			UConveyorIO.xExitBarCylinderRetract2:=0;
			iStep:=0;
		END_IF;
	END_CASE;
3:(*上料到出口*)
	CASE iStep OF
	0:(*各种初始化，能自动去3*)
		ConveyorIODown.xLoad:=0;
		ConveyorIOleft.xLoad:=0;
		ConveyorIORight.xLoad:=0;
		ConveyorIODown.xUnload:=0;
		ConveyorIOLeft.xUnload:=0;
		ConveyorIORight.xUnload:=0;
		UConveyorIO.xBatteryError:=0;
		UConveyorIO.xExitBarCylinderRetract1:=0;
		UConveyorIO.xExitBarCylinderRetract2:=0;
		ConveyorIODown.xPutInto:=0;
		ConveyorIOLeft.xPutInto:=0;
		ConveyorIORight.xPutInto:=0;
		IF m_xStep0 AND  ConveyorIODown.xEmpty THEN
			iStep:=1;
		ELSIF m_xStep0 AND NOT ConveyorIODown.xEmpty THEN
			iStep:=3;
		END_IF;	
	1:(*右顶升动作，等load*)
		IF UConveyorIO.xLiftCylinderExtendInit2 THEN
			UConveyorIO.xLiftCylinderExtend2:=0;
			UConveyorIO.xLiftCylinderRetract2:=1;
		ELSE
			UConveyorIO.xLiftCylinderExtend2:=1;
			UConveyorIO.xLiftCylinderRetract2:=0;
		END_IF;
		IF ((NOT UConveyorIO.xLiftCylinderExtendInit2 AND UConveyorIO.xLiftCylinderExtendDetect2)
			OR ( UConveyorIO.xLiftCylinderExtendInit2 AND UConveyorIO.xLiftCylinderRetractDetect2))
			AND UConveyorIO.xEntryEnable3 THEN(*有上料请求1*)
		   	ConveyorIORight.xLoad:=1;
			iStep:=2;
		END_IF;
	2:(*Load完成*)
		IF NOT ConveyorIORight.xEmpty THEN
			ConveyorIORight.xLoad:=0;
			ConveyorIODown.diDesConveyor:=ConveyorIORight.diDesConveyor;
			ConveyorIODown.xPutInto:=1;
			istep:=3;
		END_IF;
	3:(*顶升恢复等Unload，这里等有了ExitEnable再顶升，因为可能有地方需要允许了再升降，比如倍速链*)
		UConveyorIO.xExitBarCylinderRetract2:=1;
		IF  UConveyorIO.xExitEnable1 THEN(**)
			IF UConveyorIO.xLiftCylinderExtendInit2 THEN
				UConveyorIO.xLiftCylinderExtend2:=1;
				UConveyorIO.xLiftCylinderRetract2:=0;
			ELSE
				UConveyorIO.xLiftCylinderExtend2:=0;
				UConveyorIO.xLiftCylinderRetract2:=1;
			END_IF;
		END_IF;
		IF UConveyorIO.xExitEnable1 THEN(**)
			IF(( UConveyorIO.xLiftCylinderExtendInit2 AND UConveyorIO.xLiftCylinderExtendDetect2)
				OR (NOT UConveyorIO.xLiftCylinderExtendInit2 AND UConveyorIO.xLiftCylinderRetractDetect2))THEN
				ConveyorIODown.xPutInto:=0;
				iStep:=4;
			END_IF;	
		END_IF;
	4:(*Unload完成，回0*)
		IF  UConveyorIO.xExitEnable1 AND m_xExitBarDelay THEN
			ConveyorIODown.xUnload:=1;
		ELSE
			ConveyorIODown.xUnload:=0;
		END_IF;	
		IF NOT UConveyorIO.xExitEnable1 AND m_xExitBarDelay  THEN
			ConveyorIODown.xUnload:=0;
			ConveyorIOLeft.xUnload:=0;
			ConveyorIORight.xUnload:=0;
			ConveyorIODown.xPutInto:=1;
			ConveyorIOLeft.xPutInto:=1;
			ConveyorIORight.xPutInto:=1;
			UConveyorIO.xExitBarCylinderRetract1:=0;
			UConveyorIO.xExitBarCylinderRetract2:=0;
			iStep:=0;
		END_IF;
	END_CASE;
END_CASE;(*iTask*)
END_IF;(*g_xAuto那个IF*)
(*复位程序*)
IF (g_xResetSingle AND  (g_diDeviceIDSelect=ConveyorIOLeft.diDeviceID 
 	 OR g_diDeviceIDSelect=ConveyorIORight.diDeviceID
 	 OR g_diDeviceIDSelect=ConveyorIODown.diDeviceID))
	OR LDP(TRUE,UConveyorIO.xLiftCylinderExtendInit1) 
	OR LDF(TRUE,UConveyorIO.xLiftCylinderExtendInit1) 
	OR LDP(TRUE,UConveyorIO.xPutInto)  THEN
	ConveyorIODown.xPutInto:=1;
	ConveyorIOLeft.xPutInto:=1;
	ConveyorIORight.xPutInto:=1;
	iStep:=0;
END_IF;
(*手动*)
IF g_xManual  THEN
	iStep:=0;
	ConveyorIODown.xLoad:=0;
	ConveyorIOleft.xLoad:=0;
	ConveyorIORight.xLoad:=0;
	ConveyorIODown.xUnload:=0;
	ConveyorIOLeft.xUnload:=0;
	ConveyorIORight.xUnload:=0;
	ConveyorIODown.xPutInto:=0;
	ConveyorIOLeft.xPutInto:=0;
	ConveyorIORight.xPutInto:=0;
	UConveyorIO.xBatteryError:=0;
	UConveyorIO.xLiftCylinderExtend1:=UConveyorIO.xLiftCylinderExtendButton1 AND NOT UConveyorIO.xLiftCylinderRetractButton1;
	UConveyorIO.xLiftCylinderRetract1:=UConveyorIO.xLiftCylinderRetractButton1 AND NOT UConveyorIO.xLiftCylinderExtendButton1;
	UConveyorIO.xLiftCylinderExtend2:=UConveyorIO.xLiftCylinderExtendButton2 AND NOT UConveyorIO.xLiftCylinderRetractButton2;
	UConveyorIO.xLiftCylinderRetract2:=UConveyorIO.xLiftCylinderRetractButton2 AND NOT UConveyorIO.xLiftCylinderExtendButton2;
	UConveyorIO.xExitBarCylinderRetract1:=UConveyorIO.xExitBarCylinderRetractButton1;
	UConveyorIO.xExitBarCylinderRetract2:=UConveyorIO.xExitBarCylinderRetractButton2;
END_IF;	
(*气缸超时报警*)
m_tonCylinderOvertime(IN:= (UConveyorIO.xLiftCylinderExtend1 AND NOT UConveyorIO.xLiftCylinderExtendDetect1) 
 		OR  (UConveyorIO.xLiftCylinderRetract1 AND NOT UConveyorIO.xLiftCylinderRetractDetect1)
 		OR	(UConveyorIO.xLiftCylinderExtend2 AND NOT UConveyorIO.xLiftCylinderExtendDetect2) 
 		OR  (UConveyorIO.xLiftCylinderRetract2 AND NOT UConveyorIO.xLiftCylinderRetractDetect2),
 PT:= UConveyorIO.tSetOvertime ,Q:=UConveyorIO.xOvertimeAlarm ,ET:=m_tCylinderOvertimeCurrent );
END_FUNCTION_BLOCK

FUNCTION ShuttleCarCurrentPosition
VAR_INPUT
  xPosition1 : BOOL;
  xPosition2 : BOOL;
  xPosition3 : BOOL;
END_VAR
(*//计算输送车当前位置的函数*)
IF xPosition1 THEN
	ShuttleCarCurrentPosition:=1;
END_IF;
IF xPosition2 THEN
	ShuttleCarCurrentPosition:=2;
END_IF;
IF xPosition3 THEN
	ShuttleCarCurrentPosition:=3;
END_IF;
END_FUNCTION

PROGRAM 批量复制专用
SortConveyorIO30121 .i_xSortOver:=X66;
FanucRobotIO300.i_xPickOver:=X118;(-*-机器人给的取货完成-*-)
FanucRobotIO300.i_xPutOver:=X11A;(-*-机器人给的放货完成-*-)
Y3B4:=FanucRobotIO300.o_xSortStart;(-*-给机器人的开始启动-*-)
Y3A3:=FanucRobotIO300.o_xColumn[0];(-*-给机器人的行号-*-)
Y3B5:=FanucRobotIO300.o_xColumn[1];
Y3A4:=FanucRobotIO300.o_xColumn[2];
Y3B7:=FanucRobotIO300.o_xColumn[3];
Y3A6:=FanucRobotIO300.o_xRow[0];(-*-给机器人的列号-*-)
Y3A8:=FanucRobotIO300.o_xRow[1];
Y3A7:=FanucRobotIO300.o_xRow[2];
Y3A5:=FanucRobotIO300.o_xRow[3];
Y3B6:=FanucRobotIO300.o_xPutNumber[0];(-*-给机器人的放料位置-*-)
Y3A2:=FanucRobotIO300.o_xPutNumber[1];
Y3A1:=FanucRobotIO300.o_xPutNumber[2];
Y3B8:=FanucRobotIO300.o_xPutNumber[3];
Y2A1:=FanucRobotIO300.o_xCatchCylinder;
FanucRobotIO300.i_xBatteryDetect[3]:=X7F;
FanucRobotIO300.i_xBatteryDetect[2]:=XF4;
FanucRobotIO300.i_xBatteryDetect[1]:=XF6;
FanucRobotIO300.i_xBatteryDetect[0]:=XF9;
FanucRobotIO300.i_xProtect[0]:=X7E;
FanucRobotIO300.i_xProtect[1]:=XE5;
FanucRobotIO300.i_xProtect[2]:=XE4;
FanucRobotIO300.i_xProtect[3]:=XFB;

(-*-分拣排废线调用-*-)
Servo1(ServoIO:=ServoIO1 ,xAuto:=g_xAuto ,xManual:= g_xManual );
Y300:=ServoIO1.xPLCReady;
ServoIO1.xQD75Error1:=X308;					ServoIO1.xQD75Error2:=X309;		ServoIO1.xQD75Error3:=X30A;		ServoIO1.xQD75Error4:=X30B;
ServoIO1.xQD75Busy1:=X30C;				ServoIO1.xQD75Busy2:=X30D;		ServoIO1.xQD75Busy3:=X30E;		ServoIO1.xQD75Busy4:=X30F;
ServoIO1.xQD75LocateDone1:=X314;	ServoIO1.xQD75LocateDone2:=X315;	ServoIO1.xQD75LocateDone3:=X316;	ServoIO1.xQD75LocateDone4:=X317;
Y310:=ServoIO1.xQD75LocateStart1;	Y311:=ServoIO1.xQD75LocateStart2;	Y312:=ServoIO1.xQD75LocateStart3;	Y313:=ServoIO1.xQD75LocateStart4;
(-*-刹车控制，懒得单独写，就这样了-*-)
Y2CB:=ServoIO1.xQD75LocateStart1;	Y2CF:=ServoIO1.xQD75LocateStart2;	Y2D1:=ServoIO1.xQD75LocateStart3;	Y2D3:=ServoIO1.xQD75LocateStart4;
DMOV(TRUE,U30\G800,ServoIO1.diQD75CurrentPos1);(-*-当前位置-*-)	DMOV(TRUE,U30\G900,ServoIO1.diQD75CurrentPos2);(-*-当前位置-*-)
DMOV(TRUE,U30\G1000,ServoIO1.diQD75CurrentPos3);(-*-当前位置-*-)	DMOV(TRUE,U30\G1100,ServoIO1.diQD75CurrentPos4);(-*-当前位置-*-)
U30\G1502:=ServoIO1.iReset1;(-*-轴出错复位-*-)	U30\G1602:=ServoIO1.iReset2;(-*-轴出错复位-*-)
U30\G1702:=ServoIO1.iReset3;(-*-轴出错复位-*-)	U30\G1802:=ServoIO1.iReset4;(-*-轴出错复位-*-)
U30\G1500:=ServoIO1.iLocateStartNumber1;(-*-目标地址-*-)	U30\G1600:=ServoIO1.iLocateStartNumber2;(-*-目标地址-*-)
U30\G1700:=ServoIO1.iLocateStartNumber3;(-*-目标地址-*-)	U30\G1800:=ServoIO1.iLocateStartNumber4;(-*-目标地址-*-)
END_PROGRAM

FUNCTION_BLOCK Folder
VAR_IN_OUT
  FolderIO : FolderIO;
END_VAR
VAR
  m_xInitial : BOOL;
END_VAR
VAR_IN_OUT
  FolderConveyorIO : ConveyorIO;
END_VAR
VAR_GLOBAL RETAIN
  iFolderCount : INT;
END_VAR
VAR
  istep : INT;
  m_TONLoadDelay : TON;  (* 上料完成延时 *)
  m_xLoadDelay : BOOL;  (* 上料完成延时 *)
  m_tLoadDelay : TIME;  (* 上料完成延时 *)
  m_TONUpCylinderError : TON;
  m_tUpCylinderError : TIME;
  m_TONDownCylinderError : TON;
  m_tDownCylinderError : TIME;
  m_TONGrabCylinderError : TON;
  m_tGrabCylinderError : TIME;
END_VAR
(*叠盘机*)
(*初始化*)
IF NOT m_xInitial THEN
	FolderIO.i_iFloor:=3;
	FolderIO.i_tSetOvertime:=T#5S;
	
	m_xInitial:=1;
END_IF;
(*自动*)
IF g_xAuto THEN
				m_TONLoadDelay(IN:= NOT FolderConveyorIO.xEmpty,
													PT:= T#100MS,
													Q:=m_xLoadDelay,
													ET:=m_tLoadDelay);
	CASE istep OF
		0:(*各种初始化*)
			FolderConveyorIO.xLoad:=0;
			FolderConveyorIO.xUnload:=0;
			FolderConveyorIO.xPutInto:=0;
			IF FolderConveyorIO.xEmpty THEN
				istep:=1;(*空着就去1上料*)
			END_IF;	
			IF  m_xLoadDelay  THEN(*if 有料*)
				IF  FolderIO.i_xCylinderDownExtendDetect  AND FolderIO.i_xCylinderUpExtendDetect  THEN(*if 在下层*)
					IF iFolderCount=FolderIO.i_iFloor THEN(*if 是最后一次*)
						istep:=7;
					ELSE(*不是最后一次去5，是就去7*)
						istep:=5;
					END_IF;(*if 是最后一次*)	
				ELSE(*不在下层去2*)
				istep:=2;
				END_IF;	(*if 在下层*)			
			END_IF;(*if 有料*)
			
		1:(*上料*)
			IF FolderIO.i_xEntryEnable THEN
				FolderConveyorIO.xLoad:=1;
			ELSE
				FolderConveyorIO.xLoad:=0;
			END_IF;(*not Empty了等个延时*)	

			IF m_xLoadDelay  AND (iFolderCount>0 AND iFolderCount<FolderIO.i_iFloor) THEN
				istep:=2;
			ELSIF m_xLoadDelay AND iFolderCount=0 THEN(*=0表示是第一次，第一次直接抓紧上升*)
				istep:=5;	
			END_IF;	
		2:(*下降，到2层位置*)
				FolderIO.o_xCylinderUpRetract:=0;
				FolderIO.o_xCylinderUpExtend:=1;
				FolderIO.o_xCylinderDownRetract:=1;
				FolderIO.o_xCylinderDownExtend:=0;
				IF FolderIO.i_xCylinderUpExtendDetect AND FolderIO.i_xCylinderDownRetractDetect THEN
					istep:=3;
				END_IF;
		3:	(*松开夹爪*)
		
			FolderIO.o_xCylinderGrabExtend:=0;
			FolderIO.o_xCylinderGrabRetract:=1;
			IF FolderIO.i_xCylinderGrabRetractDetect THEN
				IF iFolderCount=FolderIO.i_iFloor-1 THEN
					iFolderCount:=FolderIO.i_iFloor;(*最后一次到这里就刷新计数，方便故障恢复*)
				END_IF;	
				istep:=4;
			END_IF;	
		4:(*再下降，去1层*)
				FolderIO.o_xCylinderUpRetract:=0;
				FolderIO.o_xCylinderUpExtend:=1;
				FolderIO.o_xCylinderDownRetract:=0;
				FolderIO.o_xCylinderDownExtend:=1;
				IF FolderIO.i_xCylinderDownExtendDetect  AND FolderIO.i_xCylinderUpExtendDetect  THEN
					IF iFolderCount<FolderIO.i_iFloor-1 THEN
						istep:=5;
					ELSE
						istep:=7;
					END_IF;	
				END_IF;		
		5:(*抓紧*)
			IF FolderIO.i_xCylinderDownExtendDetect  AND FolderIO.i_xCylinderUpExtendDetect  THEN
				FolderIO.o_xCylinderGrabExtend:=1;
				FolderIO.o_xCylinderGrabRetract:=0;
				IF FolderIO.i_xCylinderGrabExtendDetect THEN
					iFolderCount:=iFolderCount+1;
					istep:=6;
				END_IF;	
			END_IF;		
		6:(*上升到3层*)
			FolderIO.o_xCylinderUpRetract:=1;
			FolderIO.o_xCylinderUpExtend:=0;
			FolderIO.o_xCylinderDownRetract:=1;
			FolderIO.o_xCylinderDownExtend:=0;
			IF FolderIO.i_xCylinderDownRetractDetect AND FolderIO.i_xCylinderUpRetractDetect THEN
				FolderConveyorIO.xPutInto:=1;(*刷新成Empty的*)
				istep:=0;
			END_IF;
		7:(*下料*)	
				IF	FolderIO.i_xExitEnable AND FolderIO.i_xCylinderGrabRetractDetect	THEN(*保证不会挂到叉手*)
				FolderConveyorIO.xUnload:=1;
			ELSE
				FolderConveyorIO.xPutInto:=1;(*刷新成Empty的*)
				FolderConveyorIO.xUnload:=0;
			END_IF;	
			IF FolderConveyorIO.xEmpty THEN(*确保空了才回0，不然还在这里等Unload信号*)
				iFolderCount:=0;
				istep:=0;
			END_IF;	 
		END_CASE;
END_IF;(*g_xAuto那个*)	
(*手动控制气缸动作*)
		IF g_xManual THEN
			FolderIO.o_xCylinderGrabExtend:=	FolderIO.i_xCylinderGrabExtendButton;	
			FolderIO.o_xCylinderGrabRetract:=	FolderIO.i_xCylinderGrabRetractButton;	
			FolderIO.o_xCylinderUpExtend:=		FolderIO.i_xCylinderUpExtendButton;	
			FolderIO.o_xCylinderUpRetract:=		FolderIO.i_xCylinderUpRetractButton;	
			FolderIO.o_xCylinderDownExtend:=	FolderIO.i_xCylinderDownExtendButton;	
			FolderIO.o_xCylinderDownRetract:=	FolderIO.i_xCylinderDownRetractButton;		
		END_IF;
		
		(*气缸超时未到达报警，可能是没气儿漏气，也可能是开关坏了，或者气缸被卡住了*)
		m_TONGrabCylinderError(IN:= (FolderIO.o_xCylinderGrabExtend AND NOT FolderIO.i_xCylinderGrabExtendDetect) 
																OR  (FolderIO.o_xCylinderGrabRetract AND NOT FolderIO.i_xCylinderGrabRetractDetect) ,
															PT:= FolderIO.i_tSetOvertime ,Q:= FolderIO.o_xGrabCylinderError,ET:= m_tGrabCylinderError);
		m_TONDownCylinderError(IN:= (FolderIO.o_xCylinderDownExtend AND NOT FolderIO.i_xCylinderDownExtendDetect) 
																OR  (FolderIO.o_xCylinderDownRetract AND NOT FolderIO.i_xCylinderDownRetractDetect) ,
															PT:= FolderIO.i_tSetOvertime ,Q:= FolderIO.o_xDownCylinderError,ET:= m_tDownCylinderError);
		m_TONUpCylinderError(IN:= (FolderIO.o_xCylinderUpExtend AND NOT FolderIO.i_xCylinderUpExtendDetect) 
																OR  (FolderIO.o_xCylinderUpRetract AND NOT FolderIO.i_xCylinderUpRetractDetect) ,
															PT:= FolderIO.i_tSetOvertime ,Q:= FolderIO.o_xUpCylinderError,ET:= m_tUpCylinderError);
END_FUNCTION_BLOCK

FUNCTION_BLOCK DivideFolder
VAR_IN_OUT
  FolderIO : FolderIO;
  FolderConveyorIO : ConveyorIO;
END_VAR
VAR_GLOBAL RETAIN
  iFolderCount : INT;
END_VAR
VAR
  m_xInitial : BOOL;
  istep : INT;
  m_TONLoadDelay : TON;  (* 上料完成延时 *)
  m_xLoadDelay : BOOL;  (* 上料完成延时 *)
  m_tLoadDelay : TIME;  (* 上料完成延时 *)
  m_TONUpCylinderError : TON;
  m_tUpCylinderError : TIME;
  m_TONDownCylinderError : TON;
  m_tDownCylinderError : TIME;
  m_TONGrabCylinderError : TON;
  m_tGrabCylinderError : TIME;
END_VAR
(*叠盘机*)
(*初始化*)
IF NOT m_xInitial THEN
	FolderIO.i_iFloor:=3;
	FolderIO.i_tSetOvertime:=T#5S;
	
	m_xInitial:=1;
END_IF;
(*自动*)
IF g_xAuto THEN
	FolderIO.o_xEntryPermit:=iFolderCount=0 AND FolderConveyorIO.xEmpty;(*空了且数量为0了，才准上料*)
	m_TONLoadDelay(IN:= NOT FolderConveyorIO.xEmpty,
											PT:= T#100MS,
											Q:=m_xLoadDelay,
											ET:=m_tLoadDelay);
	CASE istep OF
		0:(*各种初始化*)
			FolderConveyorIO.xLoad:=0;
			FolderConveyorIO.xUnload:=0;
			FolderConveyorIO.xPutInto:=0;
			IF FolderConveyorIO.xEmpty THEN(*空的情况，0时上料，其他走流程*)
				IF iFolderCount=0  THEN
					istep:=1; 					
				ELSE 
					istep:=2;
				END_IF;	
			END_IF;		
			IF m_xLoadDelay THEN
				 IF FolderIO.i_xCylinderDownExtendDetect  AND FolderIO.i_xCylinderUpExtendDetect  THEN
					istep:=3;(*如果在下层执行3*)
				ELSIF FolderIO.i_xCylinderDownRetractDetect AND FolderIO.i_xCylinderUpRetractDetect THEN
					istep:=7;(*如果在上层执行下料过程*)
				 ELSE 
				 	istep:=5;(*如果在中层执行夹紧缩回流程*)
				END_IF;		
			END_IF;
		1:(*上料*)
			IF FolderIO.i_xEntryEnable THEN
				FolderConveyorIO.xLoad:=1;
			ELSE
				FolderConveyorIO.xLoad:=0;
			END_IF;(*not Empty了等个延时*)	

			IF m_xLoadDelay THEN
				iFolderCount:=FolderIO.i_iFloor;
				istep:=5;(**上料肯定是第一次才上料，所以必然去5，抓紧上升*)
			END_IF;	
		2:(*下降，到1层位置*)
				FolderIO.o_xCylinderUpRetract:=0;
				FolderIO.o_xCylinderUpExtend:=1;
				FolderIO.o_xCylinderDownRetract:=0;
				FolderIO.o_xCylinderDownExtend:=1;
				IF FolderIO.i_xCylinderDownExtendDetect AND FolderIO.i_xCylinderUpExtendDetect THEN
					istep:=3;
				END_IF;
		3:	(*松开夹爪*)
			IF FolderIO.i_xCylinderDownExtendDetect AND FolderIO.i_xCylinderUpExtendDetect THEN
				FolderIO.o_xCylinderGrabExtend:=0;
				FolderIO.o_xCylinderGrabRetract:=1;
			END_IF;
			IF FolderIO.i_xCylinderGrabRetractDetect THEN
				IF iFolderCount=1 THEN(*最后一次到这里就刷新数据，方便复位*)
					iFolderCount:=0;
				END_IF;	
				istep:=4;
			END_IF;	
		4:(*再上升到2层*)
				FolderIO.o_xCylinderUpRetract:=0;
				FolderIO.o_xCylinderUpExtend:=1;
				FolderIO.o_xCylinderDownRetract:=1;
				FolderIO.o_xCylinderDownExtend:=0;
				IF FolderIO.i_xCylinderDownRetractDetect  AND FolderIO.i_xCylinderUpExtendDetect  THEN
					IF iFolderCount=1 THEN(*最后一次到此为止，升到2层就算完成*)
						istep:=7;
					ELSE	(*其他都走正常流程*)
						istep:=5;
					END_IF;		
				END_IF;		
		5:(*抓紧*)
			IF FolderIO.i_xCylinderDownRetractDetect  AND FolderIO.i_xCylinderUpExtendDetect  THEN
				FolderIO.o_xCylinderGrabExtend:=1;
				FolderIO.o_xCylinderGrabRetract:=0;
				IF FolderIO.i_xCylinderGrabExtendDetect THEN
					istep:=6;
				END_IF;	
			END_IF;		
		6:(*上升到3层*)
			FolderIO.o_xCylinderUpRetract:=1;
			FolderIO.o_xCylinderUpExtend:=0;
			FolderIO.o_xCylinderDownRetract:=1;
			FolderIO.o_xCylinderDownExtend:=0;
			IF FolderIO.i_xCylinderDownRetractDetect AND FolderIO.i_xCylinderUpRetractDetect THEN
				FolderConveyorIO.xPutInto:=1;
				istep:=7;
			END_IF;
		7:(*下料*)	
			IF	FolderIO.i_xExitEnable	
				AND FolderIO.i_xCylinderDownExtendDetect (*通过这些保证我没有挂到叉手*)
				AND FolderIO.i_xCylinderUpExtendDetect  
				AND FolderIO.i_xCylinderGrabRetractDetect	THEN
				FolderConveyorIO.xUnload:=1;
			ELSE
				FolderConveyorIO.xPutInto:=1;
				FolderConveyorIO.xUnload:=0;
			END_IF;	
			IF FolderConveyorIO.xEmpty THEN
				IF iFolderCount>1 THEN
					iFolderCount:=iFolderCount-1;					
					istep:=2;
				ELSE
					istep:=0;
				END_IF;	
			END_IF;		
		END_CASE;
END_IF;(*g_xAuto那个*)	
(*手动控制气缸动作*)
		IF g_xManual THEN
			FolderIO.o_xCylinderGrabExtend:=	FolderIO.i_xCylinderGrabExtendButton;	
			FolderIO.o_xCylinderGrabRetract:=	FolderIO.i_xCylinderGrabRetractButton;	
			FolderIO.o_xCylinderUpExtend:=		FolderIO.i_xCylinderUpExtendButton;	
			FolderIO.o_xCylinderUpRetract:=		FolderIO.i_xCylinderUpRetractButton;	
			FolderIO.o_xCylinderDownExtend:=	FolderIO.i_xCylinderDownExtendButton;	
			FolderIO.o_xCylinderDownRetract:=	FolderIO.i_xCylinderDownRetractButton;		
		END_IF;
		
		(*气缸超时未到达报警，可能是没气儿漏气，也可能是开关坏了，或者气缸被卡住了*)
		m_TONGrabCylinderError(IN:= (FolderIO.o_xCylinderGrabExtend AND NOT FolderIO.i_xCylinderGrabExtendDetect) 
																OR  (FolderIO.o_xCylinderGrabRetract AND NOT FolderIO.i_xCylinderGrabRetractDetect) ,
															PT:= FolderIO.i_tSetOvertime ,Q:= FolderIO.o_xGrabCylinderError,ET:= m_tGrabCylinderError);
		m_TONDownCylinderError(IN:= (FolderIO.o_xCylinderDownExtend AND NOT FolderIO.i_xCylinderDownExtendDetect) 
																OR  (FolderIO.o_xCylinderDownRetract AND NOT FolderIO.i_xCylinderDownRetractDetect) ,
															PT:= FolderIO.i_tSetOvertime ,Q:= FolderIO.o_xDownCylinderError,ET:= m_tDownCylinderError);
		m_TONUpCylinderError(IN:= (FolderIO.o_xCylinderUpExtend AND NOT FolderIO.i_xCylinderUpExtendDetect) 
																OR  (FolderIO.o_xCylinderUpRetract AND NOT FolderIO.i_xCylinderUpRetractDetect) ,
															PT:= FolderIO.i_tSetOvertime ,Q:= FolderIO.o_xUpCylinderError,ET:= m_tUpCylinderError);
END_FUNCTION_BLOCK

FUNCTION_BLOCK ConveyorCommunication
VAR_IN_OUT
  ConveyorIO : ConveyorIO;
  CommunicationIO : CommunicationIO;
END_VAR
VAR_OUTPUT
  o_iErrorNub : INT;  (* 错误代码 *)
  o_xReqSuccess : BOOL;  (* 请求成功 *)
END_VAR
VAR
  m_xInitial : BOOL;  (* 初始化 *)
  o_xError : BOOL;  (* 通信数据错误 *)
END_VAR
(********************************************************************************)
(*
DB1区(PC->PLC)15个字		
"字(16位）序号
(从1开始)"			功能描述											具体参数解释
1					请求确认	"										1：复位
				 														2：读码(入库申请）成功
				 														3：取放货完成 
																		4：旋转
																		5：不旋转
																		101：条码空
																		102：条码规则校验失败
																		103：步号校验失败
																		104：无库位可用 
"
2	预留	
3	预留	
4	预留	
5	预留	
6	读写标志位	"														1：写入数据
																		2：读数据完成"
7	任务处理标志	"														１：复位
																		２：完成"
8	命令字	"
																		21-送出（任务起点与终点不同，即向下一台输送机移载）
																		22：叠盘
"
9	任务号	"															1~65535唯一任务标识"
10	目标设备号															只有送出任务才有效
11		
12	筐码后4位	
				

DB2区(PLC->PC)15个字			
"字(16位）序号
(从1开始)"	功能描述	具体参数解释	
1	请求状态	"１：复位
２：请求"	实时状态，没有时序交互
2	强制入库(预留）	"１：复位
２：强制入库"	
3	预留(叠盘数量）	只对叠盘工位有效	
4	预留		
5			
6	读写标志位	"1：写入数据
2：读数据完成"	"有交互
时序"
7	设备状态	"1:空闲
2：工作中
3:任务完成（只有目标设备才会报任务完成）
４：故障"	
8	任务号	1~65535唯一任务标识，当输送任务执行完成后，将PC下发的任务号上报	
9	筐码后4位		
10	预留		
11			
			





2018.8.3 YAO 1.0
*)
(********************************************************************************)
(*如果外部不设置，就认为没有额外条件，有料就请求*)
IF NOT m_xInitial THEN
		CommunicationIO.i_xExtraCondition:=1;
		CommunicationIO.i_xExportConveyor:=0;
		m_xInitial:=1;
END_IF;
(*//有料状态*)
IF ConveyorIO.xEmpty THEN
	CommunicationIO.o_iEmptyPLCPC:=1;
	CommunicationIO.o_iRequestPLCPC:=1;(*无料取消请求*)
ELSE
	CommunicationIO.o_iEmptyPLCPC:=2;
END_IF;

(*//请求状态*)
IF CommunicationIO.i_xExportConveyor=0 THEN(*入库段线体,有料且满足额外条件才请求*)
		IF NOT ConveyorIO.xEmpty AND CommunicationIO.i_xExtraCondition THEN
			CommunicationIO.o_iRequestPLCPC:=2;
		ELSE
			CommunicationIO.o_iRequestPLCPC:=1;
		END_IF;
ELSE(*出库段线体，有料发请求*)
		IF ConveyorIO.xEmpty AND CommunicationIO.i_xExtraCondition THEN
			CommunicationIO.o_iRequestPLCPC:=2;
		ELSE
			CommunicationIO.o_iRequestPLCPC:=1;
		END_IF;
END_IF;	
(*//请求确认*)
CASE CommunicationIO.i_iResponsPCPLC OF 
	0:;
	1:;(*//复位*)
	2:(*//读码（入库申请）成功*)
	o_xReqSuccess:=1;
	3:(*//取放货完成*)
	ConveyorIO.xPutInto:=1; 
	4:(*//旋转*)
	o_xReqSuccess:=1;
	ConveyorIO.xPutInto:=1; 
	5:(*//不旋转*)
	o_xReqSuccess:=1;
	ConveyorIO.xPutInto:=1; 
	101:(*//条码空*)
	o_iErrorNub:=101;
	o_xError:=1;
	102:(*//条码规则检验失败*)
	o_iErrorNub:=102;
	o_xError:=1;
	103:(*//步号校验失败*)
	o_iErrorNub:=103;
	o_xError:=1;
	104:(*//无库位可用*)
	o_iErrorNub:=104;
	o_xError:=1;
	105:(*//路径选择失败*)
	o_iErrorNub:=105;
	o_xError:=1;
	106:(*//控制ID错误*)
	o_iErrorNub:=106;
	o_xError:=1;
	107:(*//叠盘计数不一致*)
	o_iErrorNub:=107;
	o_xError:=1;
END_CASE;
(*IF LDP(TRUE,CommunicationIO.i_iResponsPCPLC=3
			OR CommunicationIO.i_iResponsPCPLC =4
			OR CommunicationIO.i_iResponsPCPLC =5 ) THEN
	ConveyorIO.xPutInto:=1;
END_IF;*)
IF LDP(TRUE,CommunicationIO.i_iResponsPCPLC <> 3
			AND CommunicationIO.i_iResponsPCPLC <>4
			AND CommunicationIO.i_iResponsPCPLC <>5 ) THEN
	ConveyorIO.xPutInto:=0;
END_IF;
IF CommunicationIO.i_iResponsPCPLC <> 2 
			AND CommunicationIO.i_iResponsPCPLC <>4
			AND CommunicationIO.i_iResponsPCPLC <>5 
	THEN
	o_xReqSuccess:=0;
END_IF;
IF CommunicationIO.i_iResponsPCPLC < 100 THEN
	o_iErrorNub:=0;
	o_xError:=0;
END_IF;

(*//读写标志位写入数据*)
IF ConveyorIO.diDesConveyor<>ConveyorIO.diDeviceID THEN
	IF LDP(TRUE,CommunicationIO.i_iReadWriteFlagPCPLC = 1) THEN(*标志位为1时把数据传进来*)
		ConveyorIO.iTaskID := CommunicationIO.i_iTaskIDPCPLC;
		ConveyorIO.diDesConveyor := CommunicationIO.i_diDestinationDevicePCPLC;
		ConveyorIO.iProductCategory :=CommunicationIO.i_iProductIDPCPLC;
	END_IF;
END_IF;
(*//数据校验，并返回握手信号*)
IF CommunicationIO.i_iReadWriteFlagPCPLC = 1 
			AND ConveyorIO.iTaskID<>0
			AND ConveyorIO.diDesConveyor<>0 
		  	(*AND ConveyorIO.iProductCategory<>0 *)
	THEN
	CommunicationIO.o_iReadWriteFlagPLCPC:=2;(*数据校验没问题，我们读写标志位发2*)
ELSIF CommunicationIO.i_iTaskProcessFlagPCPLC=2 THEN	(*处理标志位为2时，返回一个2*)
	CommunicationIO.o_iReadWriteFlagPLCPC:=2;(*他发任务处理完成，我们需要把读写标志位给2*)
ELSE
	CommunicationIO.o_iReadWriteFlagPLCPC:=1;
END_IF;

(*//数据校验*)
IF CommunicationIO.i_iReadWriteFlagPCPLC = 1 
			AND (ConveyorIO.iTaskID<>0
			OR ConveyorIO.diDesConveyor<>	0 )
			(*OR ConveyorIO.iProductCategory<>0) *)
	THEN
	o_iErrorNub:=50;(*//任务数据不完整*)
END_IF;
(*//设备状态*)
IF ConveyorIO.diDesConveyor = ConveyorIO.diDeviceID THEN(*//目标地址=当前地址，表示是终点设备*)
		IF  (LDP(TRUE,NOT ConveyorIO.xEmpty AND CommunicationIO.i_xExtraCondition) (*有料的上升沿报完成*)
					OR (g_diDeviceIDSelect=ConveyorIO.diDeviceID AND g_xInsertTask))(*点插入任务，也报一次完成*)
			THEN
			CommunicationIO.o_iDeviceStatusPLCPC:=3;(*//任务完成*)
			CommunicationIO.o_iProductIDPLCPC:=ConveyorIO.iProductCategory;(*//条码后四位上传*)
			CommunicationIO.o_iTaskIDPLCPC:=ConveyorIO.iTaskID;(*//任务号上传*)
			CommunicationIO.o_iRequestPLCPC:=2;(*发送入库请求*)
		ELSIF  LDP(TRUE,CommunicationIO.i_iTaskProcessFlagPCPLC=1)	THEN	(*上位机给完成信号，就复位信号*)
			CommunicationIO.o_iDeviceStatusPLCPC:=1;
			CommunicationIO.o_iProductIDPLCPC:=0;(*//条码号复位*)
			CommunicationIO.o_iTaskIDPLCPC:=0;(*//任务号复位*)
		END_IF;	
ELSIF 	ConveyorIO.diDesConveyor <>ConveyorIO.diDeviceID AND ConveyorIO.xEmpty THEN(*非终点设备，无料时复位*)
	CommunicationIO.o_iDeviceStatusPLCPC:=1;
ELSIF ConveyorIO.xBusy THEN
	CommunicationIO.o_iDeviceStatusPLCPC:=2;(*//工作中*)
ELSIF ConveyorIO.xError THEN
	CommunicationIO.o_iDeviceStatusPLCPC:=4;(*//故障*)	
END_IF;
IF NOT g_xAuto THEN(*关自动全部复位*)
	CommunicationIO.o_iDeviceStatusPLCPC:=0;
	CommunicationIO.o_iEmptyPLCPC:=0;
	CommunicationIO.o_iFolderNumberPLCPC:=0;
	CommunicationIO.o_iForceInportPLCPC:=0;
	CommunicationIO.o_iProductIDPLCPC:=0;
	CommunicationIO.o_iReadWriteFlagPLCPC:=0;
	CommunicationIO.o_iRequestPLCPC:=0;
	CommunicationIO.o_iTaskIDPLCPC:=0;
END_IF;
END_FUNCTION_BLOCK

FUNCTION_BLOCK FanucRobot
VAR_IN_OUT
  FanucRobotIO : FanucRobotIO;
END_VAR
VAR
  m_iSNO : INT;
  m_xPNSPass : BOOL;  (* 收到程序号 *)
  m_tonStartDelay : TON;  (* 启动延时 *)
  m_xStartDelay : BOOL;
  m_tStartDelayCurrentTime : TIME;
END_VAR
;
END_FUNCTION_BLOCK

FUNCTION_BLOCK SortCommunication
VAR
  m_iStep : INT;
END_VAR
VAR_IN_OUT
  ConveyorIO : ConveyorIO;
  SortCommunicationIO : SortCommunicationIO;
END_VAR
VAR
  m_iCoordinateX : INT;
  m_iCoordinateY : INT;
END_VAR
VAR_IN_OUT
  FanucRobotIO : FanucRobotIO;
END_VAR
VAR_OUTPUT
  o_iErrorNub : INT;
END_VAR
VAR
  ii : INT;
END_VAR
VAR CONSTANT
  ROW_NUB : INT := 8;  (* 每排的数量 *)
END_VAR
VAR
  m_xEno : BOOL;
  m_TONPutover : TON;  (* 放货完成滤波 *)
  m_xPutover : BOOL;  (* 放货完成滤波 *)
  m_tPutover : TIME;  (* 放货完成滤波 *)
  m_iCheck : INT;  (* 校验字 *)
END_VAR
VAR_IN_OUT
  ServoIO : ServoIO;  (* QD75 *)
END_VAR
(*********************************************************)
(*
DB1区(PC->PLC)100个字		
"字(16位）序号
(从1开始)"	功能描述	具体参数解释
1	应答	"1：复位
2：读码成功(参数写入完成)
101：条码空
102：条码规则校验失败
103：步号校验失败"
2	任务处理完成	"1：复位
2：处理完成"
3	"电芯状态，
128个电芯"	一个字代表两个电芯状态，1：合格，2,3,4:NG 

DB2区(PLC->PC)10个字		
"字(16位）序号
(从1开始)"	功能描述	具体参数解释
请求	"1：无板
2：请求分拣
"
分拣完成	"1：复位
2：挑选完成
3：撤销
"
跟机器人通信13个输出，2个输入
						13个输出分别是：4个表示行，4个表示列，4个表示不良信息，1个启动信号
						2个输入分别是：抓料完成，放料完成		

*)
(*********************************************************)
IF g_xAuto THEN
	(*——这里临时改一下，暂时人工挑选,所以需要分拣完成按钮——*)	
		IF LDP(TRUE,SortCommunicationIO.i_xSortOver)THEN
			m_iStep:=4;
		END_IF;(**)
		(*夹紧气缸控制*)
		FanucRobotIO.o_xCatchCylinder:=NOT  ConveyorIO.xEmpty AND NOT SortCommunicationIO.o_xSortDone;
		
(*——以上是暂时人工分拣的，以后删掉——*)
	CASE m_iStep OF
		0:(*//初始化*)
		SortCommunicationIO.o_iRequestPLCPC:=1;
		SortCommunicationIO.o_iSortDonePLCPC:=1;
		ii:=0;
		SortCommunicationIO.o_xSortDone:=0;
		m_iStep:=1;
		
		1:(*发送框码的扫码请求*)
		IF ConveyorIO.xEmpty THEN
			SortCommunicationIO.o_iRequestPLCPC:=1;
		ELSE
			SortCommunicationIO.o_iRequestPLCPC:=2;(*发2表示有料了，他就会扫码*)
		END_IF;
		(*//请求确认*)
		IF SortCommunicationIO.o_iRequestPLCPC=2 (*加个条件，免得无脑跳Step2*)
					AND  FanucRobotIO.i_xRobotForbidden THEN(*这里其实是NOT Forbidden才对，等机器人调好再改回来*)
			CASE SortCommunicationIO.i_iResponsPCPLC OF 
			0:;
			1:;(*//复位*)
			2:(*//读码（入库申请）成功*)
				m_iStep:=2;
				ii:=0;
				m_iCoordinateX:=1;(*//框码扫码成功后把坐标改为1,1*)
				m_iCoordinateY:=1;
			3:(*//取放货完成*)
				ConveyorIO.xPutInto:=1; 
			4:(*//旋转*)
				;
			5:(*//不旋转*)
				;
			101:(*//条码空*)
				o_iErrorNub:=101;
			102:(*//条码规则检验失败*)
				o_iErrorNub:=102;
			103:(*//步号校验失败*)
				o_iErrorNub:=103;
			104:(*//无库位可用*)
				o_iErrorNub:=104;
			END_CASE;
		END_IF;	
		
		2:(*//料框位置抓取*)		
		IF ii=129 THEN(*129表示所有有问题的都抓完了*)
			m_iStep:=4;
		ELSIF ii>0 AND ii<129 AND m_iCheck<>0 
					AND NOT FanucRobotIO.i_xBatteryDetect[0]
					AND NOT FanucRobotIO.i_xBatteryDetect[1]
					AND NOT FanucRobotIO.i_xBatteryDetect[2]
					AND NOT FanucRobotIO.i_xBatteryDetect[3](*4个电池位没料*)
					 (*有不良品*)THEN
			FanucRobotIO.o_xSortStart:=1;(*//从料框取料*)
			FanucRobotIO.o_xColumn[3]:=m_iCoordinateX/8=1;(*XY的偏移量计算在末尾*)
			FanucRobotIO.o_xColumn[2]:=(m_iCoordinateX MOD 8)/4=1;
			FanucRobotIO.o_xColumn[1]:=(m_iCoordinateX MOD 4)/2=1;
			FanucRobotIO.o_xColumn[0]:=(m_iCoordinateX MOD 2)/1=1;
			FanucRobotIO.o_xRow[3]:=m_iCoordinateY/8=1;			
			FanucRobotIO.o_xRow[2]:=(m_iCoordinateY MOD 8)/4=1;
			FanucRobotIO.o_xRow[1]:=(m_iCoordinateY MOD 4)/2=1;
			FanucRobotIO.o_xRow[0]:=(m_iCoordinateY MOD 2)/1=1;
			CASE SortCommunicationIO.i_arriBatteryStatus[ii] OF
			0:(*0表示OCV2的不良品，视为阻值错误处理*)
					FanucRobotIO.o_xPutNumber[1]:=1;					
			1:(*合格*)
					;
			2:(*容量不足*)
					FanucRobotIO.o_xPutNumber[0]:=1;	
			3:(*电压不足*)
					FanucRobotIO.o_xPutNumber[1]:=1;	
			4:(*阻值错误*)
					FanucRobotIO.o_xPutNumber[2]:=1;	
			5:(*电压过高*)
					FanucRobotIO.o_xPutNumber[3]:=1;	
			END_CASE;
		END_IF;
		IF FanucRobotIO.i_xPickOver THEN(*//抓取动作完成*)
			m_iStep:=3;
		END_IF;
	
		3:(*//放入下料皮带线*)
			FanucRobotIO.o_xSortStart:=0;(*//从料框取料*)
			FanucRobotIO.o_xColumn[3]:=0;(*XY的偏移量计算在末尾*)
			FanucRobotIO.o_xColumn[2]:=0;
			FanucRobotIO.o_xColumn[1]:=0;
			FanucRobotIO.o_xColumn[0]:=0;
			FanucRobotIO.o_xRow[3]:=0;
			FanucRobotIO.o_xRow[2]:=0;
			FanucRobotIO.o_xRow[1]:=0;
			FanucRobotIO.o_xRow[0]:=0;	
		IF FanucRobotIO.i_xPutOver THEN(*//抓取动作完成*)
			(*这个得放货完成在复位，方便step2给*)
			FanucRobotIO.o_xPutNumber[0]:=0;
			FanucRobotIO.o_xPutNumber[1]:=0;
			FanucRobotIO.o_xPutNumber[2]:=0;
			FanucRobotIO.o_xPutNumber[3]:=0;
		END_IF;
		SET(LDP(TRUE,FanucRobotIO.o_xPutNumber[0]=0) AND NOT FanucRobotIO.i_xProtect[0] AND FanucRobotIO.i_xBatteryDetect[0], ServoIO.xBackHome4);
		SET(LDP(TRUE,FanucRobotIO.o_xPutNumber[1]=0) AND NOT FanucRobotIO.i_xProtect[1] AND FanucRobotIO.i_xBatteryDetect[1], ServoIO.xBackHome3);
		SET(LDP(TRUE,FanucRobotIO.o_xPutNumber[2]=0) AND NOT FanucRobotIO.i_xProtect[2] AND FanucRobotIO.i_xBatteryDetect[2] , ServoIO.xBackHome2 );				
		SET(LDP(TRUE,FanucRobotIO.o_xPutNumber[3]=0) AND NOT FanucRobotIO.i_xProtect[3] AND FanucRobotIO.i_xBatteryDetect[3] , ServoIO.xBackHome1 );
		m_TONPutover(IN:=NOT FanucRobotIO.i_xBatteryDetect[0] AND NOT FanucRobotIO.i_xBatteryDetect[1]  AND NOT FanucRobotIO.i_xBatteryDetect[2] AND NOT FanucRobotIO.i_xBatteryDetect[3] 
												AND FanucRobotIO.o_xPutNumber[0]=0 AND FanucRobotIO.o_xPutNumber[1]=0 AND FanucRobotIO.o_xPutNumber[2]=0 AND FanucRobotIO.o_xPutNumber[3]=0,
										PT:= t#100MS ,
										Q:= m_xPutover,
										ET:= m_tPutover);
	IF LDP(TRUE,m_xPutover) THEN
			m_iStep:=2;
		END_IF;								
4:
		(*4复位所有数据*)
			FanucRobotIO.o_xSortStart:=0;(*//从料框取料*)
			FanucRobotIO.o_xColumn[3]:=0;(*XY的偏移量计算在末尾*)
			FanucRobotIO.o_xColumn[2]:=0;
			FanucRobotIO.o_xColumn[1]:=0;
			FanucRobotIO.o_xColumn[0]:=0;
			FanucRobotIO.o_xRow[3]:=0;
			FanucRobotIO.o_xRow[2]:=0;
			FanucRobotIO.o_xRow[1]:=0;
			FanucRobotIO.o_xRow[0]:=0;	
			FanucRobotIO.o_xPutNumber[0]:=0;
			FanucRobotIO.o_xPutNumber[1]:=0;
			FanucRobotIO.o_xPutNumber[2]:=0;
			FanucRobotIO.o_xPutNumber[3]:=0;

		IF  NOT SortCommunicationIO.o_xSortDone  THEN(*这里表示只给一下2*)
				SortCommunicationIO.o_iSortDonePLCPC:=2;
				SortCommunicationIO.o_xSortDone:=1;
		END_IF;		
		IF SortCommunicationIO.i_iSortDoneAknPCPLC =2 THEN
			SortCommunicationIO.o_iSortDonePLCPC:=1;
			m_iCoordinateX:=1;
			m_iCoordinateY:=1;
		END_IF;
	END_CASE;			
		IF ConveyorIO.xEmpty THEN
				m_iStep:=0;
		END_IF;

	m_iCheck:=	SortCommunicationIO.i_arriBatteryStatus[5]+
							SortCommunicationIO.i_arriBatteryStatus[1]+
							SortCommunicationIO.i_arriBatteryStatus[2]+
							SortCommunicationIO.i_arriBatteryStatus[3]+
							SortCommunicationIO.i_arriBatteryStatus[4];(*连续5个电池都是0，说明这框电池没数据，就不分拣*)
	IF LDP(TRUE,m_iStep=2 AND SortCommunicationIO.i_iInfoWriteDone=2 AND m_iCheck<>0) THEN(*判断哪个地方是有问题的*)
		FOR ii:=ii+1 TO 128 BY 1 DO
			IF SortCommunicationIO.i_arriBatteryStatus[ii]<>1 AND SortCommunicationIO.i_arriBatteryStatus[ii]<>5THEN
				m_iCoordinateX:=((ii-1)/ROW_NUB);
				m_iCoordinateY:=2*((ii-1)MOD ROW_NUB)+((m_iCoordinateX+1) MOD 2);(*把上位机给的编号值对应到二维的偏移上*)(*后面这个意思奇数排+1，偶数排不加*)
				EXIT;
			END_IF;
		END_FOR;
	END_IF;
END_IF;(*g_xauto*)	
IF  g_diDeviceIDSelect=ConveyorIO.diDeviceID AND g_xResetSingle THEN(*复位线体时，同时复位步数和请求，重新来一遍*)
	m_iStep:=0;
END_IF;	
IF  NOT g_xAuto THEN
		SortCommunicationIO.o_iRequestPLCPC:=0;
		SortCommunicationIO.o_iSortDonePLCPC:=0;
END_IF;
END_FUNCTION_BLOCK

PROGRAM START
IF g_xReset THEN
	SM50:=1;
	ELSE
	SM50:=0;
END_IF;
CASE g_iState OF
	0: (*手动*)
	g_xManual:=1;
	g_xAuto:=0;	
	g_xStackLampAmber:=1;
	g_xStackLampGreen:=0;
	g_xRemoteAuto:=0;
	g_xAutoLamp:=0;
	1:(*自动*)
	g_xManual:=0;
	g_xAuto:=1;
	g_xStackLampGreen:=1;
	g_xStackLampAmber:=0;
	g_xRemoteAuto:=0;
	g_xAutoLamp:=1;
	2:	(*远程自动*)
	g_xRemoteAuto:=1;
	g_xStackLampGreen:=1;
	g_xStackLampAmber:=0;
	g_xAuto:=0;
	g_xManual:=0;
	g_xAutoLamp:=0;
	3:(*自动未启动*)
	g_xRemoteAuto:=1;
	g_xStackLampGreen:=SM412;
	g_xStackLampAmber:=0;
	g_xAuto:=0;
	g_xManual:=0;	
	g_xAutoLamp:=0;
END_CASE;

IF g_xAutoSwitch AND g_xAutoStart  THEN  
	g_iState:=1;
END_IF;

IF g_xAutoSwitch AND (g_iState<>1 OR NOT g_xStop)  THEN  
	g_iState:=3;
END_IF;

g_xStackLampRed:=g_xAlarm AND SM412;
g_xBuzzer:=g_xAlarm AND SM412 AND NOT g_xMute;

IF NOT g_xAlarm THEN
	g_xMute:=0;
END_IF;

IF NOT g_xAutoSwitch  OR g_xEStop=0 THEN 
	g_iState:=0;
END_IF;
IF g_xRemoteAutoStart THEN
	g_iState:=2;
END_IF;
IF g_xPause AND SM412 THEN
	g_xStackLampGreen:=0;
	g_xStackLampAmber:=0;
END_IF;
END_PROGRAM

FUNCTION_BLOCK Servo
VAR_IN_OUT
  ServoIO : ServoIO;  (* 伺服IO *)
  xAuto : BOOL;  (* 自动 *)
  xManual : BOOL;  (* 手动 *)
END_VAR
VAR
  iStep : INT;  (* 流程步骤号 *)
  g_xLocate1 : BOOL;  (* 无意义 *)
END_VAR
(*PLC要给QD75就绪信号*)
ServoIO.xPLCReady:=1;
(*当前位置读取*)
DMOVP(SM412,ServoIO.diQD75CurrentPos1,ServoIO.diQD75LastPos1);(*记录1S前的位置，和现在的位置比较，判断是否需要重新启动*)
DMOVP(SM412,ServoIO.diQD75CurrentPos2,ServoIO.diQD75LastPos2);(*记录1S前的位置，和现在的位置比较，判断是否需要重新启动*)
DMOVP(SM412,ServoIO.diQD75CurrentPos3,ServoIO.diQD75LastPos3);(*记录1S前的位置，和现在的位置比较，判断是否需要重新启动*)
DMOVP(SM412,ServoIO.diQD75CurrentPos4,ServoIO.diQD75LastPos4);(*记录1S前的位置，和现在的位置比较，判断是否需要重新启动*)
IF 		 (ServoIO.xQD75LocateStart1 AND ServoIO.diQD75CurrentPos1=ServoIO.diQD75LastPos1 )
	 OR (ServoIO.xQD75LocateStart2 AND ServoIO.diQD75CurrentPos2=ServoIO.diQD75LastPos2 )
 	OR (ServoIO.xQD75LocateStart3 AND ServoIO.diQD75CurrentPos3=ServoIO.diQD75LastPos3 )
 	OR (ServoIO.xQD75LocateStart4 AND ServoIO.diQD75CurrentPos4=ServoIO.diQD75LastPos4 )
	  THEN
				ServoIO.xResetServo:=1;
ELSE
				ServoIO.xResetServo:=0;
END_IF;	
IF LDP(TRUE,ServoIO.xResetServo) THEN
	ServoIO.iReset1:=1;(*1轴复位*)
	ServoIO.iReset2:=1;(*2轴复位*)
	ServoIO.iReset3:=1;(*3轴复位*)
	ServoIO.iReset4:=1;(*4轴复位*)	
END_IF;
(*1轴回原点*)
IF ServoIO.xBackHome1 AND NOT ServoIO.xQD75LocateDone1 THEN
	ServoIO.iLocateStartNumber1:=9001;
	ServoIO.xQD75LocateStart1:=NOT ServoIO.xResetServo AND NOT ServoIO.xQD75LocateDone1;
ELSE
	ServoIO.xQD75LocateStart1:=0;
END_IF;	
	RST(LDP(TRUE,ServoIO.diQD75CurrentPos1=0) , ServoIO.xBackHome1);
(*2轴回原点*)
IF ServoIO.xBackHome2 AND NOT ServoIO.xQD75LocateDone2 THEN
	ServoIO.iLocateStartNumber2:=9001;
	ServoIO.xQD75LocateStart2:=NOT ServoIO.xResetServo AND NOT ServoIO.xQD75LocateDone2 ;
ELSE
	ServoIO.xQD75LocateStart2:=0;
END_IF;	
	RST(LDP(TRUE,ServoIO.diQD75CurrentPos2=0) ,ServoIO.xBackHome2);		
(*3轴回原点*)
IF ServoIO.xBackHome3 AND NOT ServoIO.xQD75LocateDone3 THEN
	ServoIO.iLocateStartNumber3:=9001;
	ServoIO.xQD75LocateStart3:=NOT ServoIO.xResetServo AND NOT ServoIO.xQD75LocateDone3 ;
ELSE
	ServoIO.xQD75LocateStart3:=0;
END_IF;	
	RST(LDP(TRUE,ServoIO.diQD75CurrentPos3=0) ,ServoIO.xBackHome3);	
(*4轴回原点*)
IF ServoIO.xBackHome4 AND NOT ServoIO.xQD75LocateDone4 THEN
	ServoIO.iLocateStartNumber4:=9001;
	ServoIO.xQD75LocateStart4:=NOT ServoIO.xResetServo AND NOT ServoIO.xQD75LocateDone4 ;
ELSE
	ServoIO.xQD75LocateStart4:=0;
END_IF;	
	RST(LDP(TRUE,ServoIO.diQD75CurrentPos4=0) ,ServoIO.xBackHome4);
END_FUNCTION_BLOCK
